(* Logix 5000 project; controller MV vendor 1 type 14 code 217 rev 31.11; software revision 31.00; part 13 of 53 *)
(* tags used below, declared in another part *)
   BH_Draindown_ON : DINT;
   CWD : CHECKWORD_FLAGS;
   Dummy : BOOL;
   FVHRCH202 : PlantItem;   // Valve FVHRCH202
   FVHRLTX02_IP : PlantItem;   // Effluent Tank Level Transmitter
   IGI_TestBit : BOOL;
   MC_CH2_CIP_BYPASS_Conditions : BOOL;
   MC_CH2_CIP_BYPASS_DrainConditions : BOOL;
   MC_CH2_CIP_YST_Scb_Bypass : BOOL;
   MC_CH2_DRAIN : PlantItem;   // CH2_DRAIN
   MC_CH2_LF1 : PlantItem;   // CH2_LF1
   MC_CH2_PR1 : PlantItem;   // CH2_PR1
   MC_CIP_CH2_String_OK : BOOL;
   MC_CIP_EFFTank_Start_Lvl_Ok : BOOL;
   MC_copy_how_many : DINT;
   MC_data_file_value_to_move : DINT;
   MC_from_data_file : DINT;
   MC_from_data_offset : DINT;
   MC_N10 : INT[255];   // SETTINGS
   MC_N100 : INT[255];   // C1_PLC Channel 1 PLC data
   MC_N101 : INT[255];   // CH1 PC>PLC Channel 1 PC to PLC
   MC_N102 : INT[255];   // CH1 PROG Channel 1 CIP progra m
   MC_N103 : INT[255];   // CH1 ITEMS Chwd.nos.of items to be checked for Chan nel 1
   MC_N104 : INT[255];   // CH1 REPORT Channel 1 CIP report file
   MC_N108 : INT[255];   // CH1 VDATA Channel 1 CIP progra m validation data
   MC_N112 : INT[255];   // FVR DATA Data read from FV ro uting PLC
   MC_N113 : INT[255];   // MVR DATA Data read from MV ro uting PLC
   MC_N114 : INT[255];   // YP DATA
   MC_N120 : INT[255];   // C2 PLC Channel 2 PLC data
   MC_N121 : INT[255];   // CH2 PC>PLC Channel 2 PC to PLC
   MC_N122 : INT[255];   // CH2 PROG Channel 2 CIP progra m
   MC_N123 : INT[255];   // CH2 ITEMS Chwd.nos.of items to be checked for Chan nel 2
   MC_N124 : INT[255];   // CH2 REPORT Channel 2 CIP report file
   MC_N128 : INT[255];   // CH2 VDATA Channel 2 CIP progra m validation data
   MC_N160 : INT[255];   // P40 CHECK
   MC_N161 : INT[255];   // P41 CHECK
   MC_N162 : INT[255];   // P42 CHECK
   MC_N163 : INT[255];   // P43 CHECK
   MC_N164 : INT[255];   // P44 CHECK
   MC_N165 : INT[255];   // P45 CHECK
   MC_N166 : INT[255];   // P46 CHECK
   MC_N167 : INT[255];   // Original N File From SLC, No Description Available
   MC_N20 : INT[255];   // P1 PRESS Control block and da ta for P1 pressure P ID loop
   MC_N200 : INT[255];   // CHK_WORK Plant item fault che cking work area
   MC_N201 : INT[255];   // P1 CHECK CIP program 1 plant item check list
   MC_N202 : INT[255];   // P2 CHECK CIP program 2 plant item check list
   MC_N203 : INT[255];   // P3 CHECK CIP program 3 plant item check list
   MC_N204 : INT[255];   // P4 CHECK CIP program 4 plant item check list
   MC_N205 : INT[255];   // P5 CHECK CIP program 5 plant item check list
   MC_N206 : INT[255];   // P6 CHECK CIP program 6 plant item check list
   MC_N207 : INT[255];   // P7 CHECK CIP program 7 plant item check list
   MC_N208 : INT[255];   // P8 CHECK CIP program 8 plant item check list
   MC_N209 : INT[255];   // P9 CHECK CIP program 9 plant item check list
   MC_N21 : INT[255];   // P1 FLOW Control block and da ta for P1 flowrate P ID loop
   MC_N210 : INT[255];   // P10 CHECK CIP program 10 plant item check list
   MC_N211 : INT[255];   // P11 CHECK CIP program 11 plant item check list
   MC_N212 : INT[255];   // P12 CHECK CIP program 12 plant item check list
   MC_N213 : INT[255];   // P13 CHECK CIP program 13 plant item check list
   MC_N214 : INT[255];   // P14 CHECK CIP program 14 plant item check list
   MC_N215 : INT[255];   // P15 CHECK CIP program 15 plant item check list
   MC_N216 : INT[255];   // P16 CHECK CIP program 16 plant item check list
   MC_N217 : INT[255];   // P17 CHECK CIP program 17 plant item check list
   MC_N218 : INT[255];   // P18 CHECK CIP program 18 plant item check list
   MC_N219 : INT[255];   // P19 CHECK CIP program 19 plant item check list
   MC_N22 : INT[255];   // P2 PRESS Control block and da ta for P2 pressure P ID loop
   MC_N220 : INT[255];   // P20 CHECK CIP program 20 plant item check list
   MC_N221 : INT[255];   // P21 CHECK CIP program 21 plant item check list
   MC_N222 : INT[255];   // P22 CHECK CIP program 22 plant item check list
   MC_N223 : INT[255];   // P23 CHECK CIP program 23 plant item check list
   MC_N224 : INT[255];   // P24 CHECK CIP program 24 plant item check list
   MC_N23 : INT[255];   // P2 FLOW Control block and da ta for P2 flowrate P ID loop
   MC_N7 : INT[255];   // INTEGER
   MC_N80 : INT[255];   // SRV1_PLC Detergent tank 1 ser vice PLC data
   MC_N81 : INT[255];   // SV1_PC Detergent tank 1 ser vice PC to PLC data
   MC_N82 : INT[255];   // SV1 ITEMS Chwd.nos.of items to be checked for DT1 service
   MC_N90 : INT[255];   // SV2_PLC Detergent tank 2 ser vice PLC data
   MC_N91 : INT[255];   // SV2_PC Detergent tank 2 ser vice PC to PLC data
   MC_N92 : INT[255];   // SV2 ITEMS Chwd.nos.of items to be checked for DT2 service
   MC_T125 : TIMER[255];   // CH2 TIMERS Channel 2 timers
   MC_T4 : TIMER[255];   // TIMER
   MC_to_data_file : DINT;
   MC_to_data_offset : DINT;
(* MC_Common, continued *)

ROUTINE MC_CH2_PRERN_131   (* ladder *)
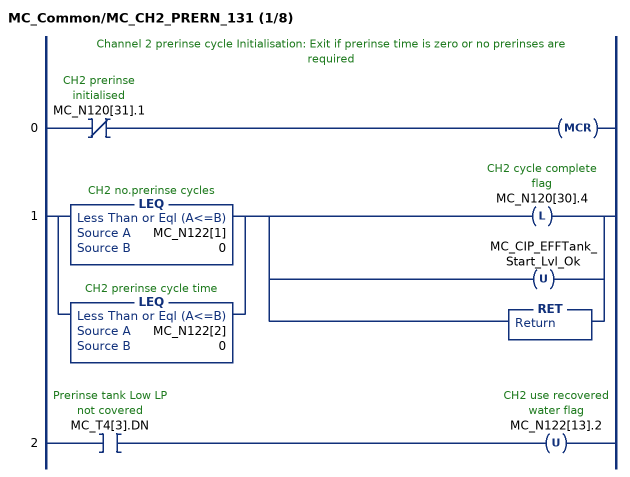
   // Channel 2 prerinse cycle Initialisation: Exit if prerinse time is zero or no prerinses are required
   0: XIO(MC_N120[31].1)MCR();
   1: [LEQ(MC_N122[1],0) ,LEQ(MC_N122[2],0) ][OTL(MC_N120[30].4) ,OTU(MC_CIP_EFFTank_Start_Lvl_Ok) ,RET() ];
   2: XIC(MC_T4[3].DN)OTU(MC_N122[13].2);
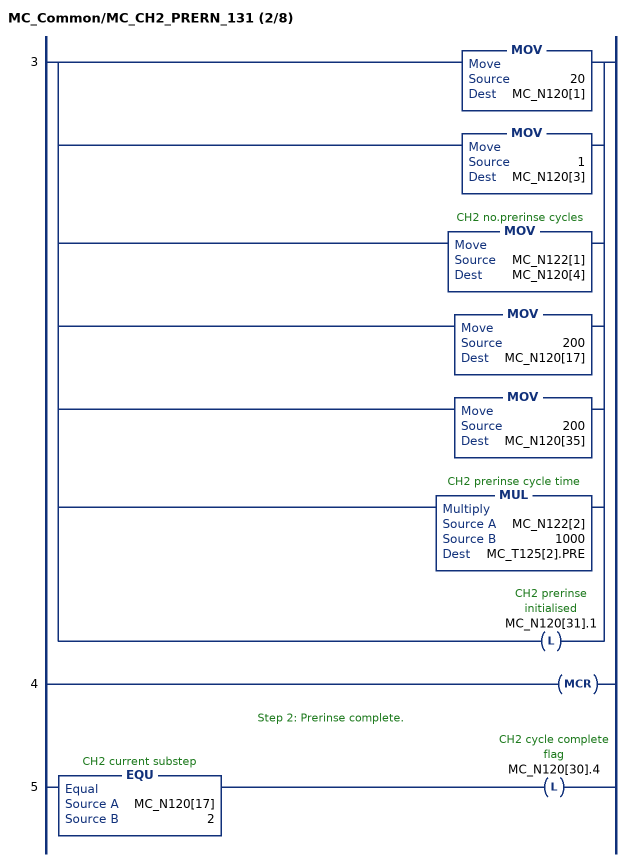
   3: [MOV(20,MC_N120[1]) ,MOV(1,MC_N120[3]) ,MOV(MC_N122[1],MC_N120[4]) ,MOV(200,MC_N120[17]) ,MOV(200,MC_N120[35]) ,MUL(MC_N122[2],1000,MC_T125[2].PRE) ,OTL(MC_N120[31].1) ];
   4: MCR();
   // Step 2: Prerinse complete.
   5: EQU(MC_N120[17],2)OTL(MC_N120[30].4);
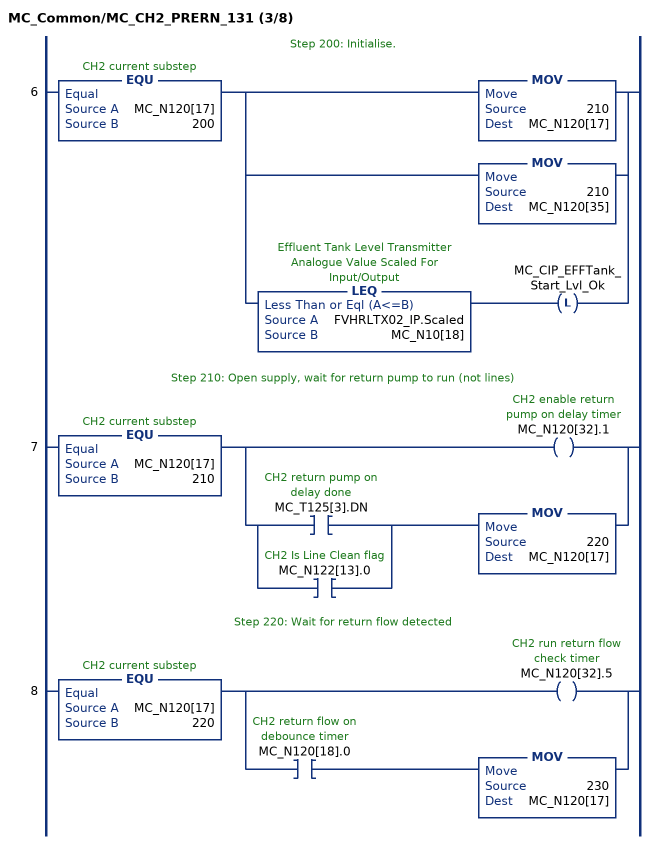
   // Step 200: Initialise.
   6: EQU(MC_N120[17],200)[MOV(210,MC_N120[17]) ,MOV(210,MC_N120[35]) ,LEQ(FVHRLTX02_IP.Scaled,MC_N10[18]) OTL(MC_CIP_EFFTank_Start_Lvl_Ok) ];
   // Step 210: Open supply, wait for return pump to run (not lines)
   7: EQU(MC_N120[17],210)[OTE(MC_N120[32].1) ,[XIC(MC_T125[3].DN) ,XIC(MC_N122[13].0) ] MOV(220,MC_N120[17]) ];
   // Step 220: Wait for return flow detected
   8: EQU(MC_N120[17],220)[OTE(MC_N120[32].5) ,XIC(MC_N120[18].0) MOV(230,MC_N120[17]) ];
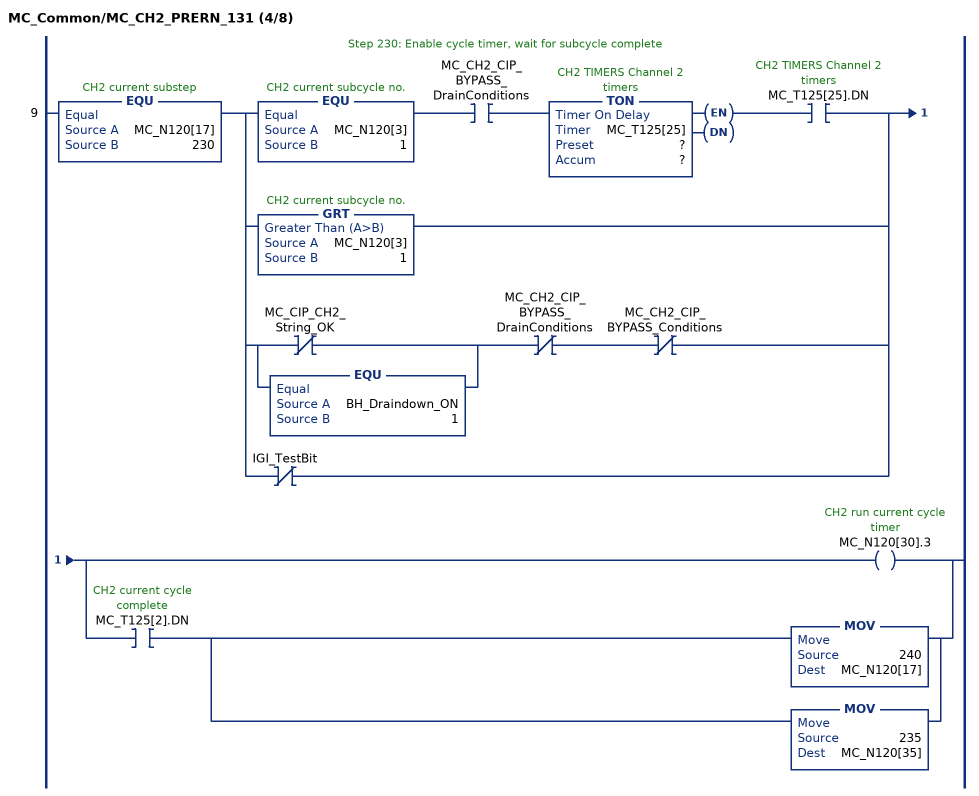
   // Step 230: Enable cycle timer, wait for subcycle complete
   9: EQU(MC_N120[17],230)[EQU(MC_N120[3],1) XIC(MC_CH2_CIP_BYPASS_DrainConditions) TON(MC_T125[25],?,?) XIC(MC_T125[25].DN) ,GRT(MC_N120[3],1) ,[XIO(MC_CIP_CH2_String_OK) ,EQU(BH_Draindown_ON,1) ] XIO(MC_CH2_CIP_BYPASS_DrainConditions) XIO(MC_CH2_CIP_BYPASS_Conditions) ,XIO(IGI_TestBit) ][OTE(MC_N120[30].3) ,XIC(MC_T125[2].DN) [MOV(240,MC_N120[17]) ,MOV(235,MC_N120[35]) ] ];
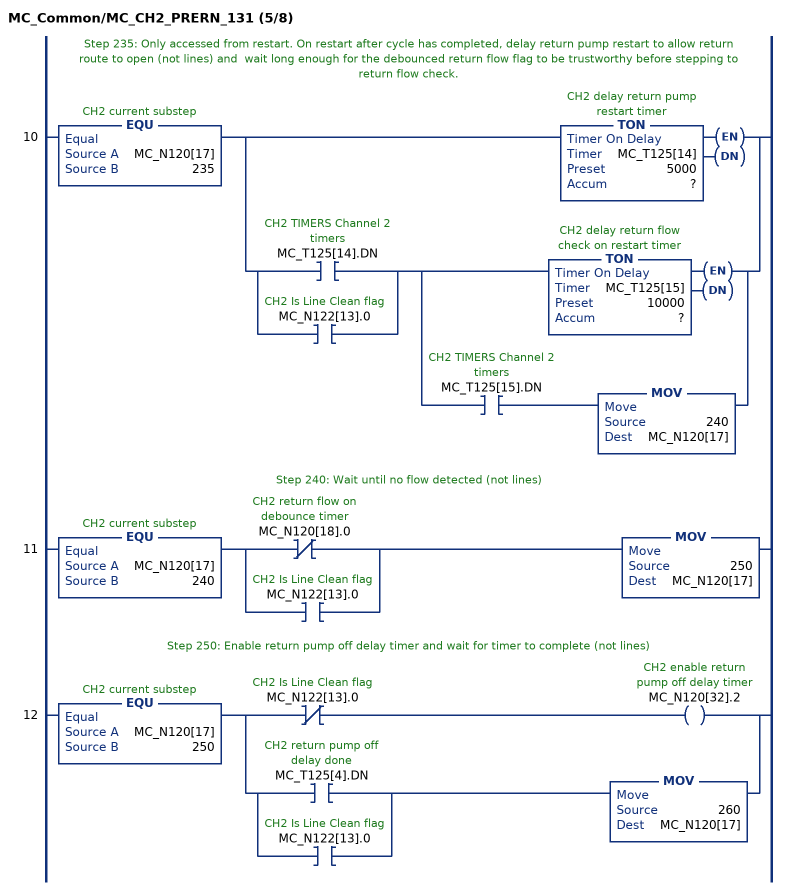
   // Step 235: Only accessed from restart. On restart after cycle has completed, delay return pump restart to allow return route to open (not lines) and  wait long enough for the debounced return flow flag to be trustworthy before stepping to return flow check.
   10: EQU(MC_N120[17],235)[TON(MC_T125[14],?,?) ,[XIC(MC_T125[14].DN) ,XIC(MC_N122[13].0) ] [TON(MC_T125[15],?,?) ,XIC(MC_T125[15].DN) MOV(240,MC_N120[17]) ] ];
   // Step 240: Wait until no flow detected (not lines)
   11: EQU(MC_N120[17],240)[XIO(MC_N120[18].0) ,XIC(MC_N122[13].0) ]MOV(250,MC_N120[17]);
   // Step 250: Enable return pump off delay timer and wait for timer to complete (not lines)
   12: EQU(MC_N120[17],250)[XIO(MC_N122[13].0) OTE(MC_N120[32].2) ,[XIC(MC_T125[4].DN) ,XIC(MC_N122[13].0) ] MOV(260,MC_N120[17]) ];
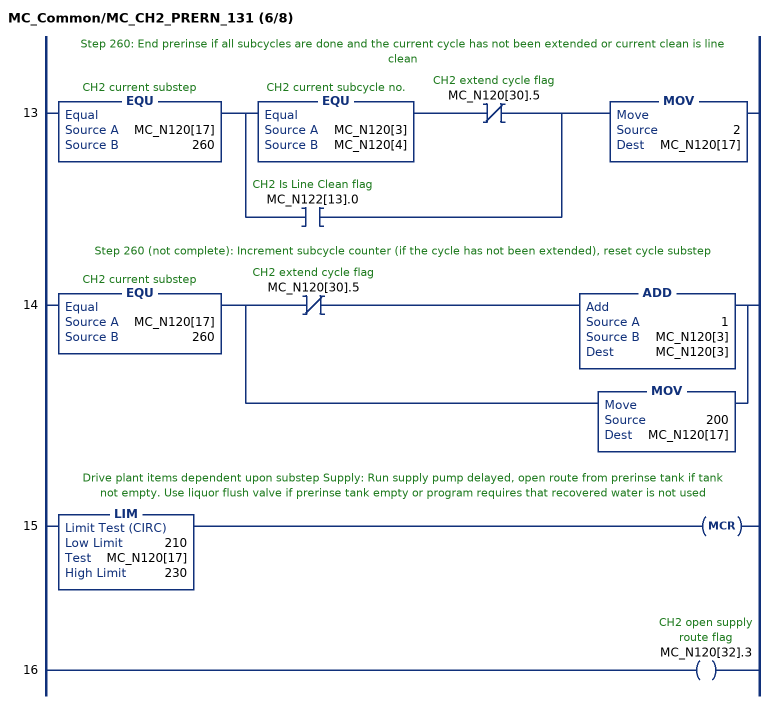
   // Step 260: End prerinse if all subcycles are done and the current cycle has not been extended or current clean is line clean
   13: EQU(MC_N120[17],260)[EQU(MC_N120[3],MC_N120[4]) XIO(MC_N120[30].5) ,XIC(MC_N122[13].0) ]MOV(2,MC_N120[17]);
   // Step 260 (not complete): Increment subcycle counter (if the cycle has not been extended), reset cycle substep
   14: EQU(MC_N120[17],260)[XIO(MC_N120[30].5) ADD(1,MC_N120[3],MC_N120[3]) ,MOV(200,MC_N120[17]) ];
   // Drive plant items dependent upon substep Supply: Run supply pump delayed, open route from prerinse tank if tank not empty. Use liquor flush valve if prerinse tank empty or program requires that recovered water is not used
   15: LIM(210,MC_N120[17],230)MCR();
   16: OTE(MC_N120[32].3);
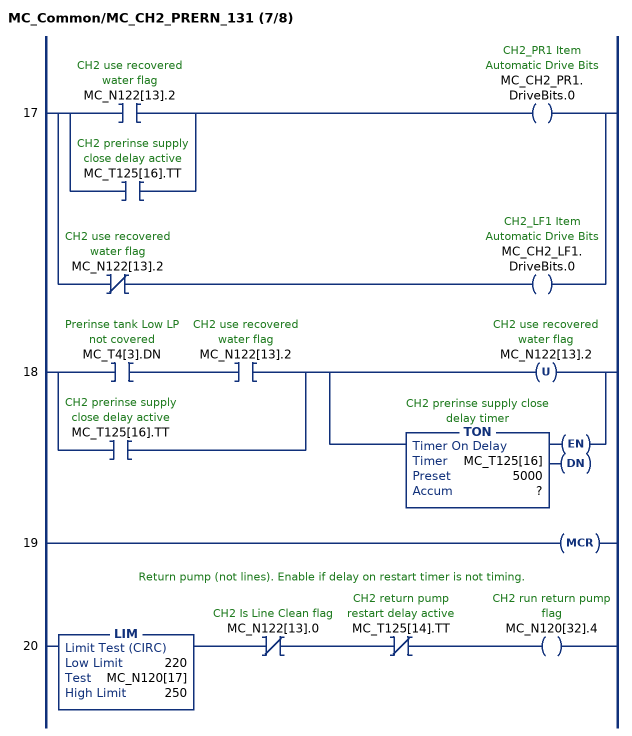
   17: [[XIC(MC_N122[13].2) ,XIC(MC_T125[16].TT) ] OTE(MC_CH2_PR1.DriveBits.0) ,XIO(MC_N122[13].2) OTE(MC_CH2_LF1.DriveBits.0) ];
   18: [XIC(MC_T4[3].DN) XIC(MC_N122[13].2) ,XIC(MC_T125[16].TT) ][OTU(MC_N122[13].2) ,TON(MC_T125[16],?,?) ];
   19: MCR();
   // Return pump (not lines). Enable if delay on restart timer is not timing.
   20: LIM(220,MC_N120[17],250)XIO(MC_N122[13].0)XIO(MC_T125[14].TT)OTE(MC_N120[32].4);
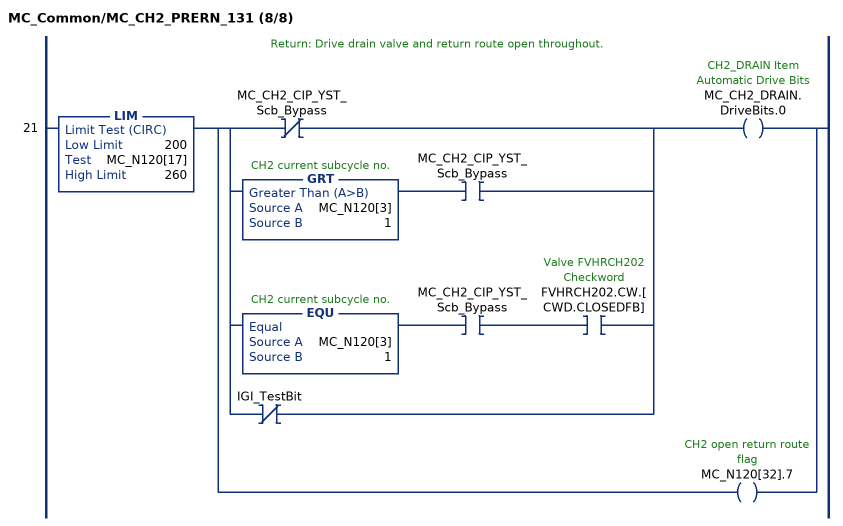
   // Return: Drive drain valve and return route open throughout.
   21: LIM(200,MC_N120[17],260)[[XIO(MC_CH2_CIP_YST_Scb_Bypass) ,GRT(MC_N120[3],1) XIC(MC_CH2_CIP_YST_Scb_Bypass) ,EQU(MC_N120[3],1) XIC(MC_CH2_CIP_YST_Scb_Bypass) XIC(FVHRCH202.CW.[CWD.CLOSEDFB]) ,XIO(IGI_TestBit) ] OTE(MC_CH2_DRAIN.DriveBits.0) ,OTE(MC_N120[32].7) ];
END_ROUTINE

ROUTINE MC_CH2_REPORT_124   (* ladder *)
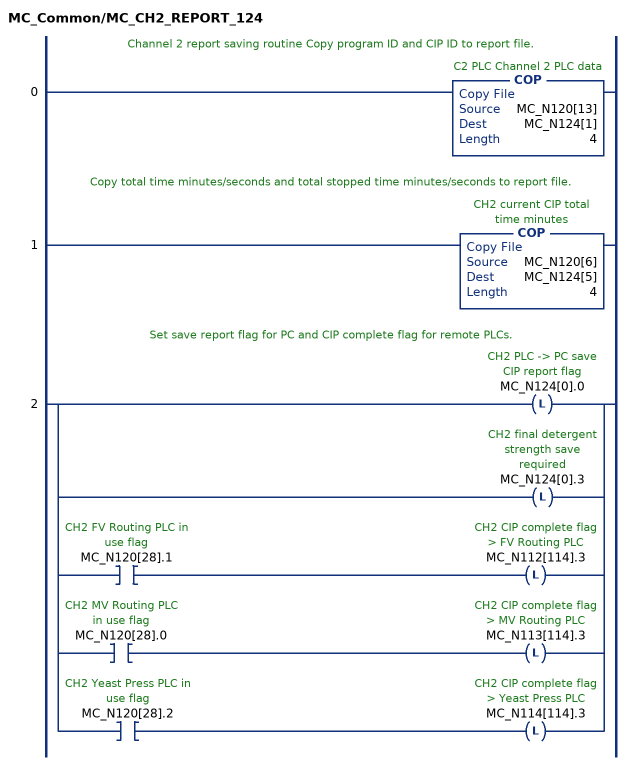
   // Channel 2 report saving routine Copy program ID and CIP ID to report file.
   0: COP(MC_N120[13],MC_N124[1],4);
   // Copy total time minutes/seconds and total stopped time minutes/seconds to report file.
   1: COP(MC_N120[6],MC_N124[5],4);
   // Set save report flag for PC and CIP complete flag for remote PLCs.
   2: [OTL(MC_N124[0].0) ,OTL(MC_N124[0].3) ,XIC(MC_N120[28].1) OTL(MC_N112[114].3) ,XIC(MC_N120[28].0) OTL(MC_N113[114].3) ,XIC(MC_N120[28].2) OTL(MC_N114[114].3) ];
END_ROUTINE

ROUTINE MC_CH2_SCAV_130   (* ladder *)
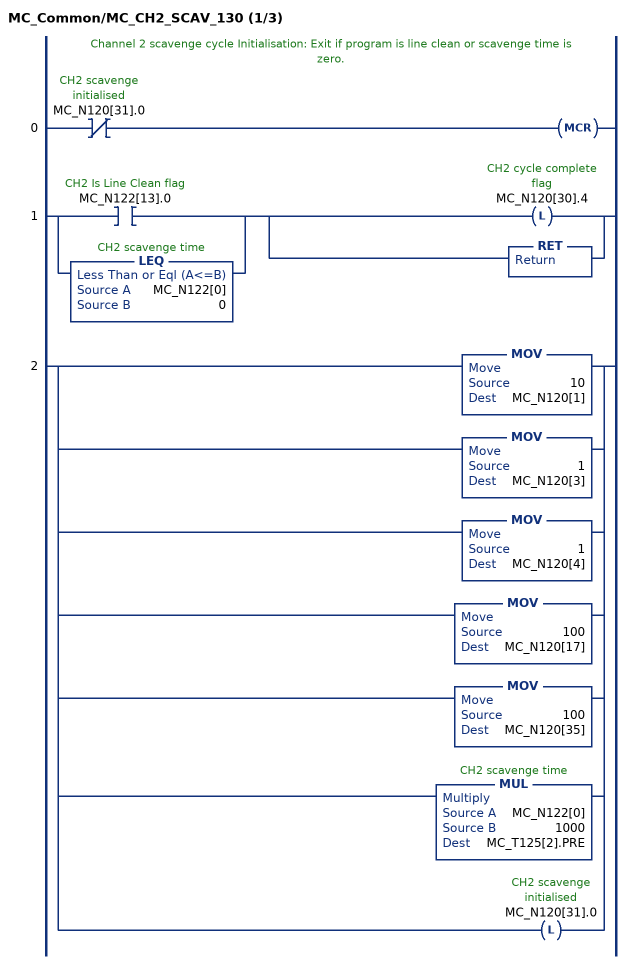
   // Channel 2 scavenge cycle Initialisation: Exit if program is line clean or scavenge time is zero.
   0: XIO(MC_N120[31].0)MCR();
   1: [XIC(MC_N122[13].0) ,LEQ(MC_N122[0],0) ][OTL(MC_N120[30].4) ,RET() ];
   2: [MOV(10,MC_N120[1]) ,MOV(1,MC_N120[3]) ,MOV(1,MC_N120[4]) ,MOV(100,MC_N120[17]) ,MOV(100,MC_N120[35]) ,MUL(MC_N122[0],1000,MC_T125[2].PRE) ,OTL(MC_N120[31].0) ];
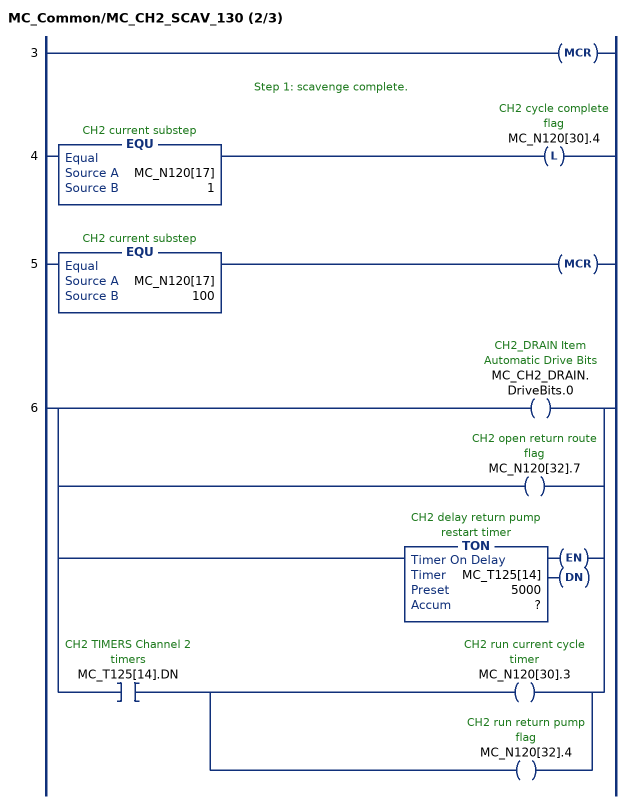
   3: MCR();
   // Step 1: scavenge complete.
   4: EQU(MC_N120[17],1)OTL(MC_N120[30].4);
   5: EQU(MC_N120[17],100)MCR();
   6: [[OTE(MC_CH2_DRAIN.DriveBits.0) ,OTE(MC_N120[32].7) ] ,[TON(MC_T125[14],?,?) ,XIC(MC_T125[14].DN) [OTE(MC_N120[30].3) ,OTE(MC_N120[32].4) ] ] ];
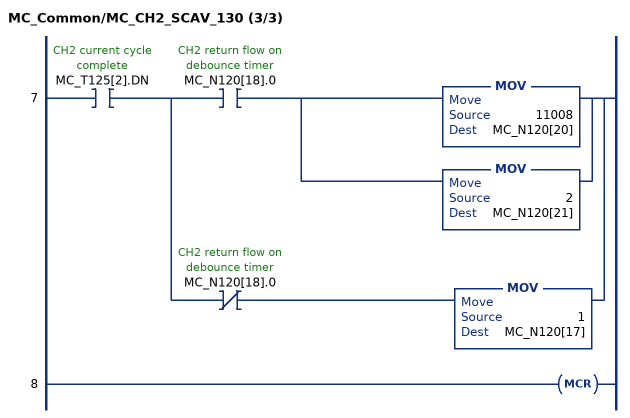
   7: XIC(MC_T125[2].DN)[XIC(MC_N120[18].0) [MOV(11008,MC_N120[20]) ,MOV(2,MC_N120[21]) ] ,XIO(MC_N120[18].0) MOV(1,MC_N120[17]) ];
   8: MCR();
END_ROUTINE

ROUTINE MC_CH2_VALID_128   (* ladder *)
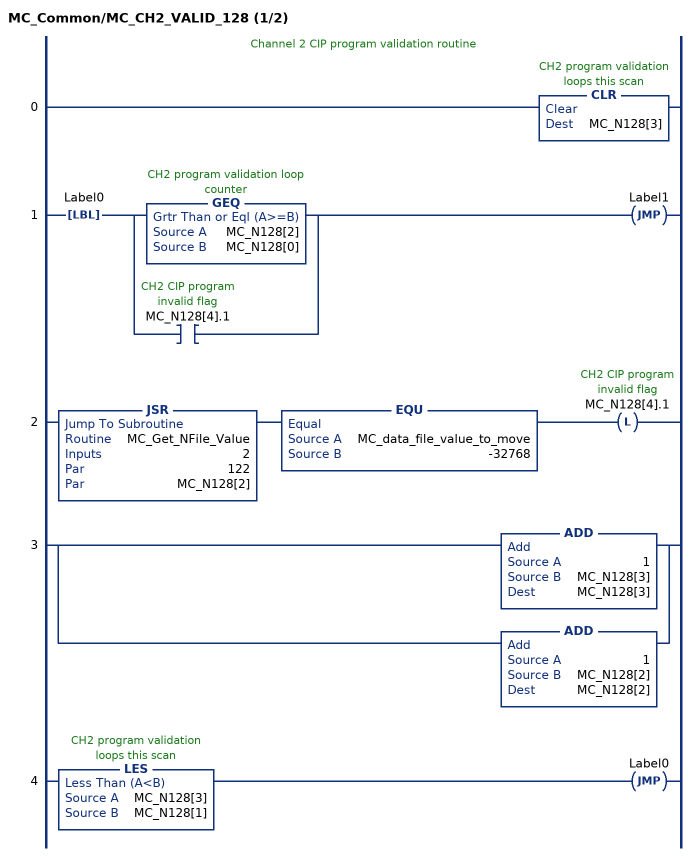
   // Channel 2 CIP program validation routine
   0: CLR(MC_N128[3]);
   1: LBL(Label0)[GEQ(MC_N128[2],MC_N128[0]) ,XIC(MC_N128[4].1) ]JMP(Label1);
   2: JSR(MC_Get_NFile_Value,2,122,MC_N128[2])EQU(MC_data_file_value_to_move,-32768)OTL(MC_N128[4].1);
   3: [ADD(1,MC_N128[3],MC_N128[3]) ,ADD(1,MC_N128[2],MC_N128[2]) ];
   4: LES(MC_N128[3],MC_N128[1])JMP(Label0);
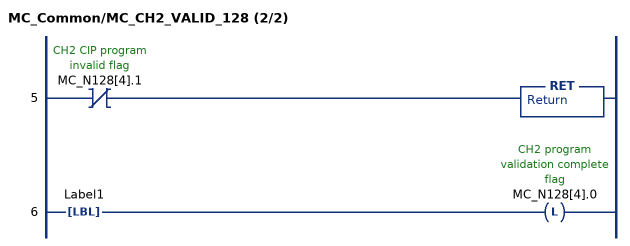
   5: XIO(MC_N128[4].1)RET();
   6: LBL(Label1)OTL(MC_N128[4].0);
END_ROUTINE

ROUTINE MC_Copy_NFile_Block   (* ladder *)
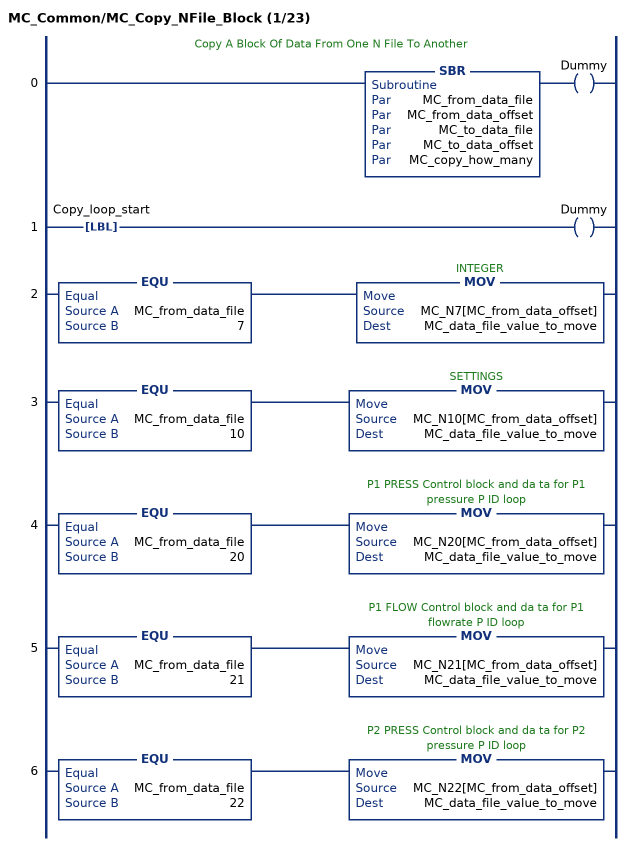
   // Copy A Block Of Data From One N File To Another
   0: SBR(MC_from_data_file,MC_from_data_offset,MC_to_data_file,MC_to_data_offset,MC_copy_how_many)OTE(Dummy);
   1: LBL(Copy_loop_start)OTE(Dummy);
   2: EQU(MC_from_data_file,7)MOV(MC_N7[MC_from_data_offset],MC_data_file_value_to_move);
   3: EQU(MC_from_data_file,10)MOV(MC_N10[MC_from_data_offset],MC_data_file_value_to_move);
   4: EQU(MC_from_data_file,20)MOV(MC_N20[MC_from_data_offset],MC_data_file_value_to_move);
   5: EQU(MC_from_data_file,21)MOV(MC_N21[MC_from_data_offset],MC_data_file_value_to_move);
   6: EQU(MC_from_data_file,22)MOV(MC_N22[MC_from_data_offset],MC_data_file_value_to_move);
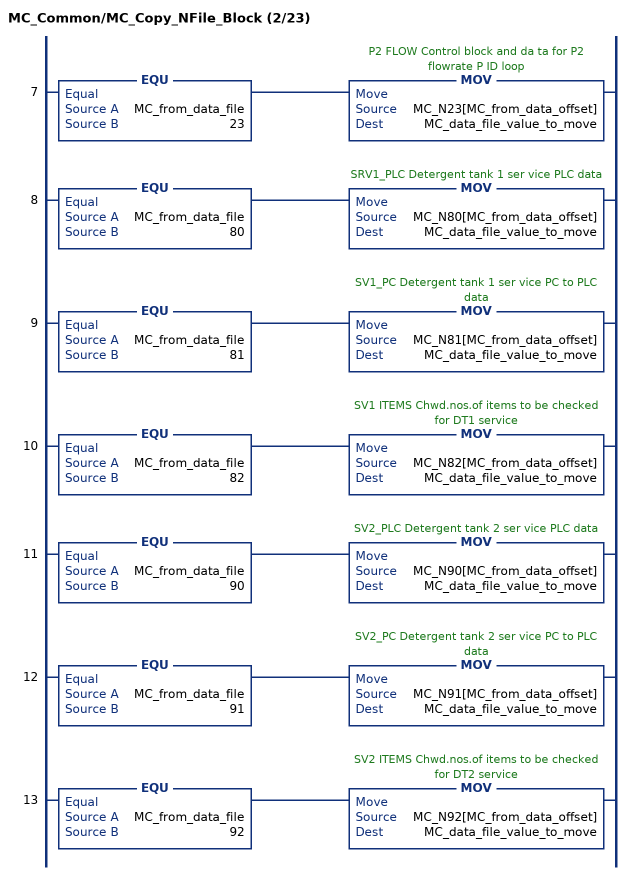
   7: EQU(MC_from_data_file,23)MOV(MC_N23[MC_from_data_offset],MC_data_file_value_to_move);
   8: EQU(MC_from_data_file,80)MOV(MC_N80[MC_from_data_offset],MC_data_file_value_to_move);
   9: EQU(MC_from_data_file,81)MOV(MC_N81[MC_from_data_offset],MC_data_file_value_to_move);
   10: EQU(MC_from_data_file,82)MOV(MC_N82[MC_from_data_offset],MC_data_file_value_to_move);
   11: EQU(MC_from_data_file,90)MOV(MC_N90[MC_from_data_offset],MC_data_file_value_to_move);
   12: EQU(MC_from_data_file,91)MOV(MC_N91[MC_from_data_offset],MC_data_file_value_to_move);
   13: EQU(MC_from_data_file,92)MOV(MC_N92[MC_from_data_offset],MC_data_file_value_to_move);
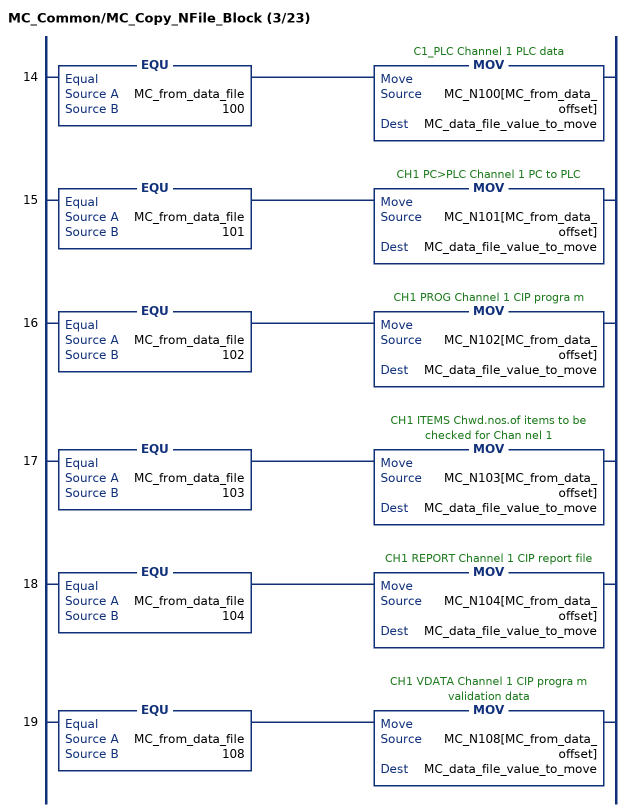
   14: EQU(MC_from_data_file,100)MOV(MC_N100[MC_from_data_offset],MC_data_file_value_to_move);
   15: EQU(MC_from_data_file,101)MOV(MC_N101[MC_from_data_offset],MC_data_file_value_to_move);
   16: EQU(MC_from_data_file,102)MOV(MC_N102[MC_from_data_offset],MC_data_file_value_to_move);
   17: EQU(MC_from_data_file,103)MOV(MC_N103[MC_from_data_offset],MC_data_file_value_to_move);
   18: EQU(MC_from_data_file,104)MOV(MC_N104[MC_from_data_offset],MC_data_file_value_to_move);
   19: EQU(MC_from_data_file,108)MOV(MC_N108[MC_from_data_offset],MC_data_file_value_to_move);
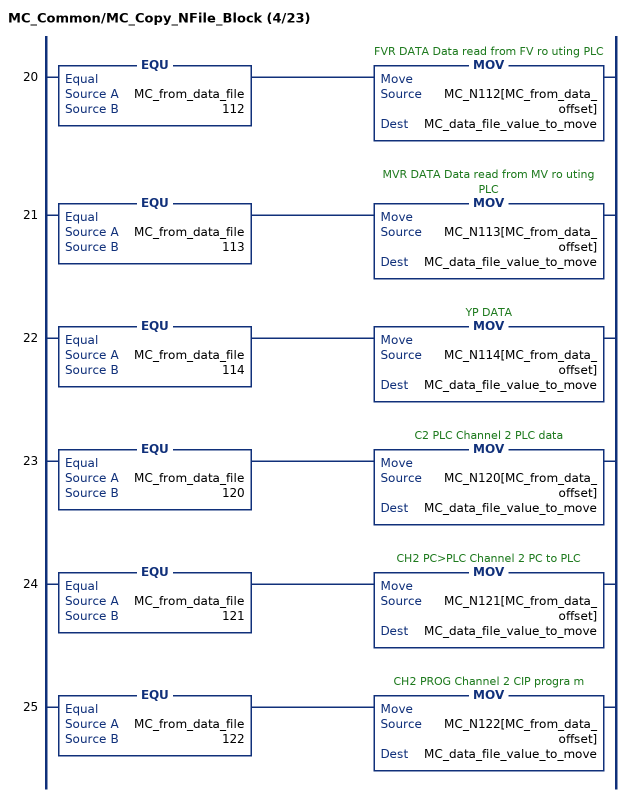
   20: EQU(MC_from_data_file,112)MOV(MC_N112[MC_from_data_offset],MC_data_file_value_to_move);
   21: EQU(MC_from_data_file,113)MOV(MC_N113[MC_from_data_offset],MC_data_file_value_to_move);
   22: EQU(MC_from_data_file,114)MOV(MC_N114[MC_from_data_offset],MC_data_file_value_to_move);
   23: EQU(MC_from_data_file,120)MOV(MC_N120[MC_from_data_offset],MC_data_file_value_to_move);
   24: EQU(MC_from_data_file,121)MOV(MC_N121[MC_from_data_offset],MC_data_file_value_to_move);
   25: EQU(MC_from_data_file,122)MOV(MC_N122[MC_from_data_offset],MC_data_file_value_to_move);
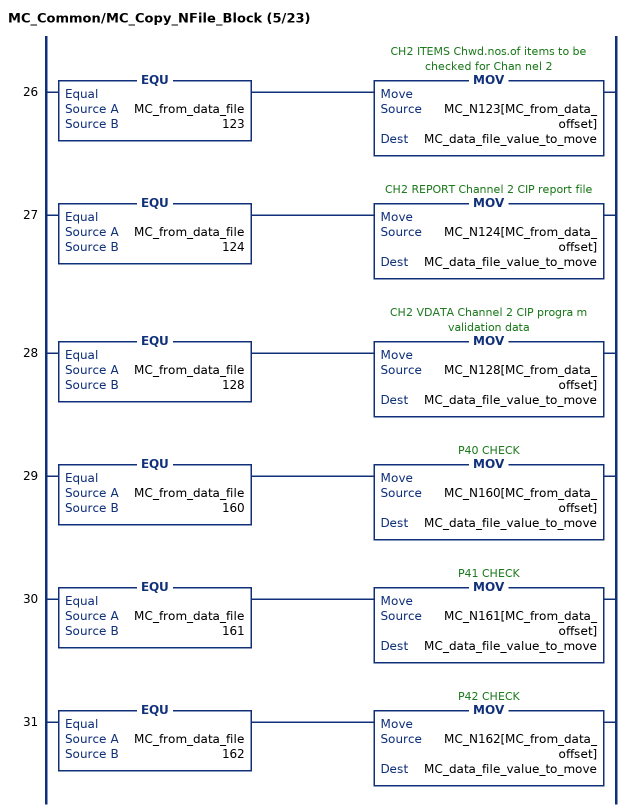
   26: EQU(MC_from_data_file,123)MOV(MC_N123[MC_from_data_offset],MC_data_file_value_to_move);
   27: EQU(MC_from_data_file,124)MOV(MC_N124[MC_from_data_offset],MC_data_file_value_to_move);
   28: EQU(MC_from_data_file,128)MOV(MC_N128[MC_from_data_offset],MC_data_file_value_to_move);
   29: EQU(MC_from_data_file,160)MOV(MC_N160[MC_from_data_offset],MC_data_file_value_to_move);
   30: EQU(MC_from_data_file,161)MOV(MC_N161[MC_from_data_offset],MC_data_file_value_to_move);
   31: EQU(MC_from_data_file,162)MOV(MC_N162[MC_from_data_offset],MC_data_file_value_to_move);
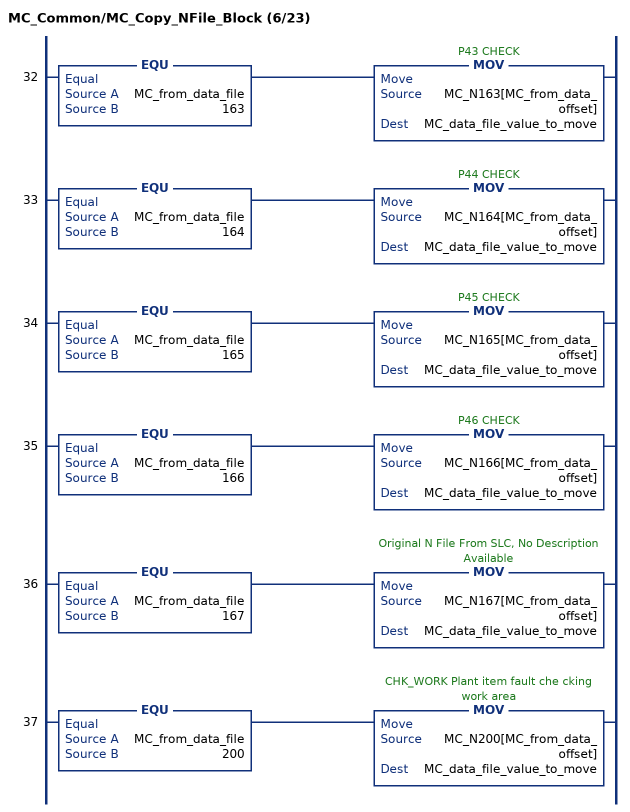
   32: EQU(MC_from_data_file,163)MOV(MC_N163[MC_from_data_offset],MC_data_file_value_to_move);
   33: EQU(MC_from_data_file,164)MOV(MC_N164[MC_from_data_offset],MC_data_file_value_to_move);
   34: EQU(MC_from_data_file,165)MOV(MC_N165[MC_from_data_offset],MC_data_file_value_to_move);
   35: EQU(MC_from_data_file,166)MOV(MC_N166[MC_from_data_offset],MC_data_file_value_to_move);
   36: EQU(MC_from_data_file,167)MOV(MC_N167[MC_from_data_offset],MC_data_file_value_to_move);
   37: EQU(MC_from_data_file,200)MOV(MC_N200[MC_from_data_offset],MC_data_file_value_to_move);
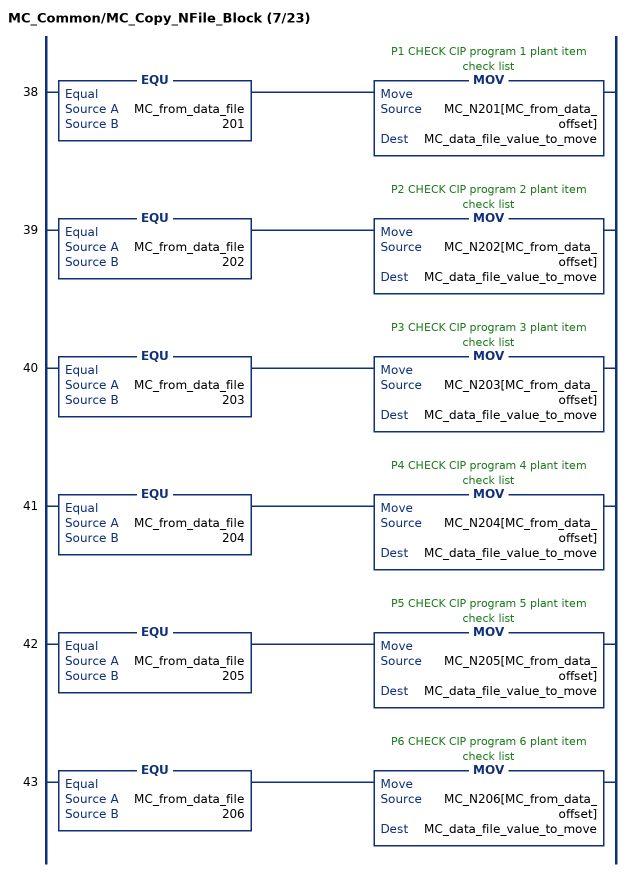
   38: EQU(MC_from_data_file,201)MOV(MC_N201[MC_from_data_offset],MC_data_file_value_to_move);
   39: EQU(MC_from_data_file,202)MOV(MC_N202[MC_from_data_offset],MC_data_file_value_to_move);
   40: EQU(MC_from_data_file,203)MOV(MC_N203[MC_from_data_offset],MC_data_file_value_to_move);
   41: EQU(MC_from_data_file,204)MOV(MC_N204[MC_from_data_offset],MC_data_file_value_to_move);
   42: EQU(MC_from_data_file,205)MOV(MC_N205[MC_from_data_offset],MC_data_file_value_to_move);
   43: EQU(MC_from_data_file,206)MOV(MC_N206[MC_from_data_offset],MC_data_file_value_to_move);
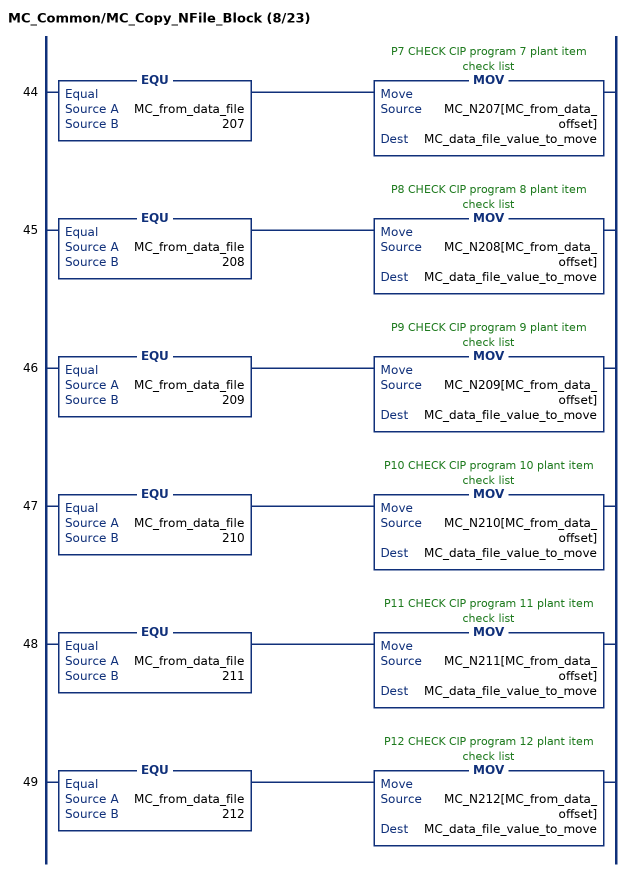
   44: EQU(MC_from_data_file,207)MOV(MC_N207[MC_from_data_offset],MC_data_file_value_to_move);
   45: EQU(MC_from_data_file,208)MOV(MC_N208[MC_from_data_offset],MC_data_file_value_to_move);
   46: EQU(MC_from_data_file,209)MOV(MC_N209[MC_from_data_offset],MC_data_file_value_to_move);
   47: EQU(MC_from_data_file,210)MOV(MC_N210[MC_from_data_offset],MC_data_file_value_to_move);
   48: EQU(MC_from_data_file,211)MOV(MC_N211[MC_from_data_offset],MC_data_file_value_to_move);
   49: EQU(MC_from_data_file,212)MOV(MC_N212[MC_from_data_offset],MC_data_file_value_to_move);
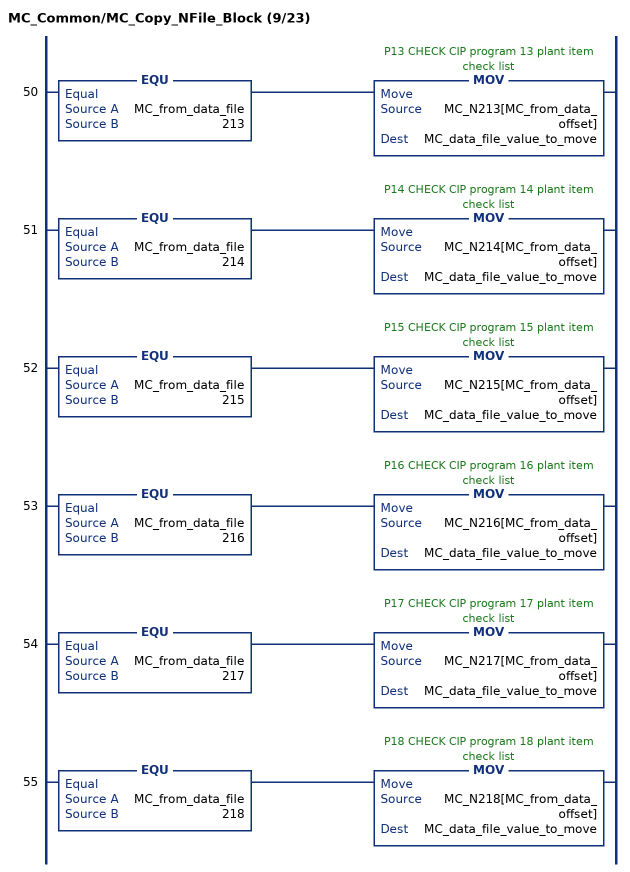
   50: EQU(MC_from_data_file,213)MOV(MC_N213[MC_from_data_offset],MC_data_file_value_to_move);
   51: EQU(MC_from_data_file,214)MOV(MC_N214[MC_from_data_offset],MC_data_file_value_to_move);
   52: EQU(MC_from_data_file,215)MOV(MC_N215[MC_from_data_offset],MC_data_file_value_to_move);
   53: EQU(MC_from_data_file,216)MOV(MC_N216[MC_from_data_offset],MC_data_file_value_to_move);
   54: EQU(MC_from_data_file,217)MOV(MC_N217[MC_from_data_offset],MC_data_file_value_to_move);
   55: EQU(MC_from_data_file,218)MOV(MC_N218[MC_from_data_offset],MC_data_file_value_to_move);
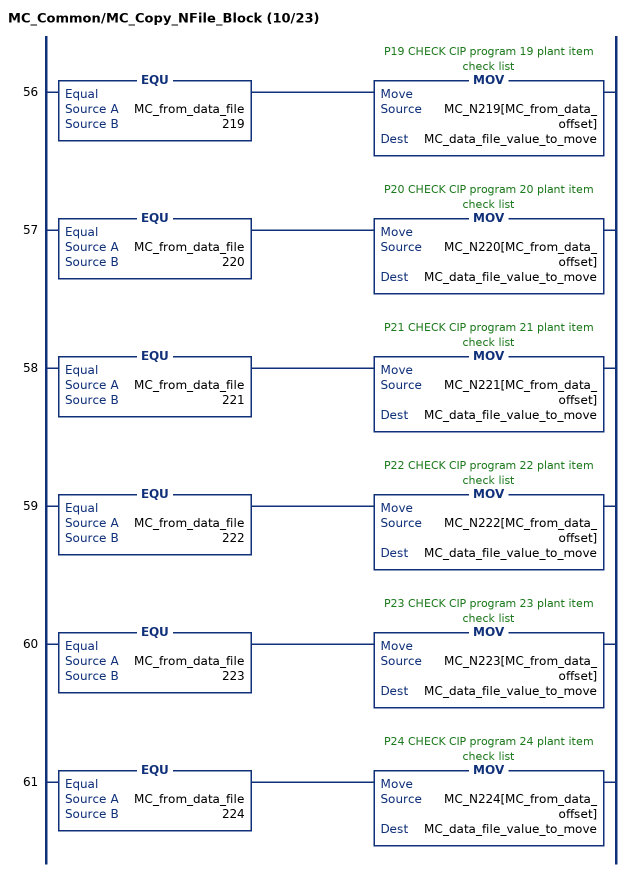
   56: EQU(MC_from_data_file,219)MOV(MC_N219[MC_from_data_offset],MC_data_file_value_to_move);
   57: EQU(MC_from_data_file,220)MOV(MC_N220[MC_from_data_offset],MC_data_file_value_to_move);
   58: EQU(MC_from_data_file,221)MOV(MC_N221[MC_from_data_offset],MC_data_file_value_to_move);
   59: EQU(MC_from_data_file,222)MOV(MC_N222[MC_from_data_offset],MC_data_file_value_to_move);
   60: EQU(MC_from_data_file,223)MOV(MC_N223[MC_from_data_offset],MC_data_file_value_to_move);
   61: EQU(MC_from_data_file,224)MOV(MC_N224[MC_from_data_offset],MC_data_file_value_to_move);
